         CALL  "FC071_CleaningPiston"
         ( IN_WithCP                := "DB704_MH_Value".Mixinghead[5].WithCleaningPiston,
           IN_Ana_CP_State          := #AnaCp_StatB,
           IN_SWUEnabled            := "DB619_State_MPart".SWU[1].SWU_released."05",
           IN_ButtonCPForward       := "DB123_MH_IO_Signals".MH[5].IN.MH_CP_forward,
           IN_ButtonCPback          := "DB123_MH_IO_Signals".MH[5].IN.MH_CP_backward,
           IN_CPForwardFromExternal := #Temp_CP_forward_external,
           IN_CPAfterShot           := "DB619_State_MPart".ShotMa[1].ShotData.CP_AfterShot,
           IN_PartshotDisabled      := "DB619_State_MPart".ShotMa[1].ShotData.ShotDisabled,
           IN_Blowing_OUT           := "DB614_MH_State".InertingMH[5].Start_Prepare_Purge_after_Shot,
           IN_CPProxSwitch          := "DB123_MH_IO_Signals".MH[5].IN.MH_APS_CleaningPiston,
           IN_SWUActive             := "DB619_State_MPart".SWU[1].Open_SWU_allone."05",
           IN_HydraulicOk           := "DB619_State_MPart".Machine[1].HydStartUp_finished,
           IN_ResetFaults           := "DB009_Faults".Faults_Reset_FKT_M1,
           IN_ControlVoltage        := "DB619_State_MPart".Operationmode[1].Controllvoltage,
           IN_OperatingModeValid    := "DB619_State_MPart".Operationmode[1].valid,
           IN_OperatingModeWithFoam := "DB619_State_MPart".Operationmode[1].Operation,
           IN_OperatingModeTestValv := "DB619_State_MPart".Operationmode[1].Test,
           IN_Lamptest              := "DB619_State_MPart".Operationmode[1].Lamptest,
           IN_ShotEnd               := "DB619_State_MPart".Cycle[1].PulsShotend,
           IN_FaultLevel_1          := "DB009_Faults".Fault_State_Grp_1_M1,
           IN_PressurizeTimeRunning := "DB619_State_MPart".Cycle[1].PressurizeTimeRuns,
           IN_ShotActive            := "DB619_State_MPart".Cycle[1].ShotRuns,
           IN_CycleRunning          := "DB619_State_MPart".Cycle[1].running,
           IN_RmpCtrlChangeTimeEnd  := "DB619_State_MPart".Cycle[1].RmpCtrlChangeTimeEnd,
           IN_StandbyTimeRunning    := "DB619_State_MPart".Cycle[1].StandByTimeRuns,
           IN_RmpCycleEnd           := "DB619_State_MPart".Cycle[1].PulseCycleEnd,
           IN_CPTimer               := "TM_RunTime_CP05",
           IN_TMCheckHomePos        := "TM_FltCPHomePos_CP05",
           Values                   := "DB704_MH_Value".Mixinghead[5].Cleaning_Piston,
           OUT_ValveCPForward       := "DB123_MH_IO_Signals".MH[5].OUT.MH.V_CP_Forward_MH,
           OUT_LampCPBack           := "DB123_MH_IO_Signals".MH[5].OUT.MH.H_CP_Back_MH,
           IO_CPIsOk                := "DB619_State_MPart".Mixinghead[1].Cleaningpiston_OK,
           IO_ReqHydrForCleaning    := "DB611_Hydraulic_State".MH_Hydraulic[1].Request_from_CP,
           IO_Status                := "DB614_MH_State".MH_CleaningPiston[5],
           IO_Fault                 := "DB824_Error_MH_CP".CPiston[5],
           IO_NewFault              := "DB009_Faults".Faultschanging_M1,
           IO_FaultLevel_1          := "DB009_Faults".Faults_FKT_Grp_1_M1,
           IO_FaultLevel_2          := "DB009_Faults".Faults_FKT_Grp_2_M1,
           IO_FaultLevel_3          := "DB009_Faults".Faults_FKT_Grp_3_M1
         );
END_REGION

REGION Network 11: Activate cleaning piston mixinghead by external signal
         A     "DB005_RS<->Extern".MC_Interface[6].Data_from_MC.CP_forward;
         =     #Temp_CP_forward_external;
END_REGION

REGION Network 12: Cleaning piston mixinghead 06
         CALL  BLKMOV
         ( SRCBLK  := "DB123_MH_IO_Signals".MH[6].IN.CleaningPistonState,
           RET_VAL := #RetValSFC,
           DSTBLK  := #AnaCp_Stat
         );

         L     #AnaCp_Stat;
         SRW   8;
         T     #AnaCp_StatB;

         CALL  "FC071_CleaningPiston"
         ( IN_WithCP                := "DB704_MH_Value".Mixinghead[6].WithCleaningPiston,
           IN_Ana_CP_State          := #AnaCp_StatB,
           IN_SWUEnabled            := "DB619_State_MPart".SWU[1].SWU_released."06",
           IN_ButtonCPForward       := "DB123_MH_IO_Signals".MH[6].IN.MH_CP_forward,
           IN_ButtonCPback          := "DB123_MH_IO_Signals".MH[6].IN.MH_CP_backward,
           IN_CPForwardFromExternal := #Temp_CP_forward_external,
           IN_CPAfterShot           := "DB619_State_MPart".ShotMa[1].ShotData.CP_AfterShot,
           IN_PartshotDisabled      := "DB619_State_MPart".ShotMa[1].ShotData.ShotDisabled,
           IN_Blowing_OUT           := "DB614_MH_State".InertingMH[6].Start_Prepare_Purge_after_Shot,
           IN_CPProxSwitch          := "DB123_MH_IO_Signals".MH[6].IN.MH_APS_CleaningPiston,
           IN_SWUActive             := "DB619_State_MPart".SWU[1].Open_SWU_allone."06",
           IN_HydraulicOk           := "DB619_State_MPart".Machine[1].HydStartUp_finished,
           IN_ResetFaults           := "DB009_Faults".Faults_Reset_FKT_M1,
           IN_ControlVoltage        := "DB619_State_MPart".Operationmode[1].Controllvoltage,
           IN_OperatingModeValid    := "DB619_State_MPart".Operationmode[1].valid,
           IN_OperatingModeWithFoam := "DB619_State_MPart".Operationmode[1].Operation,
           IN_OperatingModeTestValv := "DB619_State_MPart".Operationmode[1].Test,
           IN_Lamptest              := "DB619_State_MPart".Operationmode[1].Lamptest,
           IN_ShotEnd               := "DB619_State_MPart".Cycle[1].PulsShotend,
           IN_FaultLevel_1          := "DB009_Faults".Fault_State_Grp_1_M1,
           IN_PressurizeTimeRunning := "DB619_State_MPart".Cycle[1].PressurizeTimeRuns,
           IN_ShotActive            := "DB619_State_MPart".Cycle[1].ShotRuns,
           IN_CycleRunning          := "DB619_State_MPart".Cycle[1].running,
           IN_RmpCtrlChangeTimeEnd  := "DB619_State_MPart".Cycle[1].RmpCtrlChangeTimeEnd,
           IN_StandbyTimeRunning    := "DB619_State_MPart".Cycle[1].StandByTimeRuns,
           IN_RmpCycleEnd           := "DB619_State_MPart".Cycle[1].PulseCycleEnd,
           IN_CPTimer               := "TM_RunTime_CP06",
           IN_TMCheckHomePos        := "TM_FltCPHomePos_CP06",
           Values                   := "DB704_MH_Value".Mixinghead[6].Cleaning_Piston,
           OUT_ValveCPForward       := "DB123_MH_IO_Signals".MH[6].OUT.MH.V_CP_Forward_MH,
           OUT_LampCPBack           := "DB123_MH_IO_Signals".MH[6].OUT.MH.H_CP_Back_MH,
           IO_CPIsOk                := "DB619_State_MPart".Mixinghead[1].Cleaningpiston_OK,
           IO_ReqHydrForCleaning    := "DB611_Hydraulic_State".MH_Hydraulic[1].Request_from_CP,
           IO_Status                := "DB614_MH_State".MH_CleaningPiston[6],
           IO_Fault                 := "DB824_Error_MH_CP".CPiston[6],
           IO_NewFault              := "DB009_Faults".Faultschanging_M1,
           IO_FaultLevel_1          := "DB009_Faults".Faults_FKT_Grp_1_M1,
           IO_FaultLevel_2          := "DB009_Faults".Faults_FKT_Grp_2_M1,
           IO_FaultLevel_3          := "DB009_Faults".Faults_FKT_Grp_3_M1
         );
END_REGION

REGION Network 13: Activate cleaning piston mixinghead by external signal
         A     "DB005_RS<->Extern".MC_Interface[7].Data_from_MC.CP_forward;
         =     #Temp_CP_forward_external;
END_REGION

REGION Network 14: Cleaning piston mixinghead 07
         CALL  BLKMOV
         ( SRCBLK  := "DB123_MH_IO_Signals".MH[7].IN.CleaningPistonState,
           RET_VAL := #RetValSFC,
           DSTBLK  := #AnaCp_Stat
         );

         L     #AnaCp_Stat;
         SRW   8;
         T     #AnaCp_StatB;

         CALL  "FC071_CleaningPiston"
         ( IN_WithCP                := "DB704_MH_Value".Mixinghead[7].WithCleaningPiston,
           IN_Ana_CP_State          := #AnaCp_StatB,
           IN_SWUEnabled            := "DB619_State_MPart".SWU[1].SWU_released."07",
           IN_ButtonCPForward       := "DB123_MH_IO_Signals".MH[7].IN.MH_CP_forward,
           IN_ButtonCPback          := "DB123_MH_IO_Signals".MH[7].IN.MH_CP_backward,
           IN_CPForwardFromExternal := #Temp_CP_forward_external,
           IN_CPAfterShot           := "DB619_State_MPart".ShotMa[1].ShotData.CP_AfterShot,
           IN_PartshotDisabled      := "DB619_State_MPart".ShotMa[1].ShotData.ShotDisabled,
           IN_Blowing_OUT           := "DB614_MH_State".InertingMH[7].Start_Prepare_Purge_after_Shot,
           IN_CPProxSwitch          := "DB123_MH_IO_Signals".MH[7].IN.MH_APS_CleaningPiston,
           IN_SWUActive             := "DB619_State_MPart".SWU[1].Open_SWU_allone."07",
           IN_HydraulicOk           := "DB619_State_MPart".Machine[1].HydStartUp_finished,
           IN_ResetFaults           := "DB009_Faults".Faults_Reset_FKT_M1,
           IN_ControlVoltage        := "DB619_State_MPart".Operationmode[1].Controllvoltage,
           IN_OperatingModeValid    := "DB619_State_MPart".Operationmode[1].valid,
           IN_OperatingModeWithFoam := "DB619_State_MPart".Operationmode[1].Operation,
           IN_OperatingModeTestValv := "DB619_State_MPart".Operationmode[1].Test,
           IN_Lamptest              := "DB619_State_MPart".Operationmode[1].Lamptest,
           IN_ShotEnd               := "DB619_State_MPart".Cycle[1].PulsShotend,
           IN_FaultLevel_1          := "DB009_Faults".Fault_State_Grp_1_M1,
           IN_PressurizeTimeRunning := "DB619_State_MPart".Cycle[1].PressurizeTimeRuns,
           IN_ShotActive            := "DB619_State_MPart".Cycle[1].ShotRuns,
           IN_CycleRunning          := "DB619_State_MPart".Cycle[1].running,
           IN_RmpCtrlChangeTimeEnd  := "DB619_State_MPart".Cycle[1].RmpCtrlChangeTimeEnd,
           IN_StandbyTimeRunning    := "DB619_State_MPart".Cycle[1].StandByTimeRuns,
           IN_RmpCycleEnd           := "DB619_State_MPart".Cycle[1].PulseCycleEnd,
           IN_CPTimer               := "TM_RunTime_CP07",
           IN_TMCheckHomePos        := "TM_FltCPHomePos_CP07",
           Values                   := "DB704_MH_Value".Mixinghead[7].Cleaning_Piston,
           OUT_ValveCPForward       := "DB123_MH_IO_Signals".MH[7].OUT.MH.V_CP_Forward_MH,
           OUT_LampCPBack           := "DB123_MH_IO_Signals".MH[7].OUT.MH.H_CP_Back_MH,
           IO_CPIsOk                := "DB619_State_MPart".Mixinghead[1].Cleaningpiston_OK,
           IO_ReqHydrForCleaning    := "DB611_Hydraulic_State".MH_Hydraulic[1].Request_from_CP,
           IO_Status                := "DB614_MH_State".MH_CleaningPiston[7],
           IO_Fault                 := "DB824_Error_MH_CP".CPiston[7],
           IO_NewFault              := "DB009_Faults".Faultschanging_M1,
           IO_FaultLevel_1          := "DB009_Faults".Faults_FKT_Grp_1_M1,
           IO_FaultLevel_2          := "DB009_Faults".Faults_FKT_Grp_2_M1,
           IO_FaultLevel_3          := "DB009_Faults".Faults_FKT_Grp_3_M1
         );
END_REGION

REGION Network 15: Activate cleaning piston mixinghead by external signal
         A     "DB005_RS<->Extern".MC_Interface[8].Data_from_MC.CP_forward;
         =     #Temp_CP_forward_external;
END_REGION

REGION Network 16: Cleaning piston mixinghead 08
         CALL  BLKMOV
         ( SRCBLK  := "DB123_MH_IO_Signals".MH[8].IN.CleaningPistonState,
           RET_VAL := #RetValSFC,
           DSTBLK  := #AnaCp_Stat
         );

         L     #AnaCp_Stat;
         SRW   8;
         T     #AnaCp_StatB;

         CALL  "FC071_CleaningPiston"
         ( IN_WithCP                := "DB704_MH_Value".Mixinghead[8].WithCleaningPiston,
           IN_Ana_CP_State          := #AnaCp_StatB,
           IN_SWUEnabled            := "DB619_State_MPart".SWU[1].SWU_released."08",
           IN_ButtonCPForward       := "DB123_MH_IO_Signals".MH[8].IN.MH_CP_forward,
           IN_ButtonCPback          := "DB123_MH_IO_Signals".MH[8].IN.MH_CP_backward,
           IN_CPForwardFromExternal := #Temp_CP_forward_external,
           IN_CPAfterShot           := "DB619_State_MPart".ShotMa[1].ShotData.CP_AfterShot,
           IN_PartshotDisabled      := "DB619_State_MPart".ShotMa[1].ShotData.ShotDisabled,
           IN_Blowing_OUT           := "DB614_MH_State".InertingMH[8].Start_Prepare_Purge_after_Shot,
           IN_CPProxSwitch          := "DB123_MH_IO_Signals".MH[8].IN.MH_APS_CleaningPiston,
           IN_SWUActive             := "DB619_State_MPart".SWU[1].Open_SWU_allone."08",
           IN_HydraulicOk           := "DB619_State_MPart".Machine[1].HydStartUp_finished,
           IN_ResetFaults           := "DB009_Faults".Faults_Reset_FKT_M1,
           IN_ControlVoltage        := "DB619_State_MPart".Operationmode[1].Controllvoltage,
           IN_OperatingModeValid    := "DB619_State_MPart".Operationmode[1].valid,
           IN_OperatingModeWithFoam := "DB619_State_MPart".Operationmode[1].Operation,
           IN_OperatingModeTestValv := "DB619_State_MPart".Operationmode[1].Test,
           IN_Lamptest              := "DB619_State_MPart".Operationmode[1].Lamptest,
           IN_ShotEnd               := "DB619_State_MPart".Cycle[1].PulsShotend,
           IN_FaultLevel_1          := "DB009_Faults".Fault_State_Grp_1_M1,
           IN_PressurizeTimeRunning := "DB619_State_MPart".Cycle[1].PressurizeTimeRuns,
           IN_ShotActive            := "DB619_State_MPart".Cycle[1].ShotRuns,
           IN_CycleRunning          := "DB619_State_MPart".Cycle[1].running,
           IN_RmpCtrlChangeTimeEnd  := "DB619_State_MPart".Cycle[1].RmpCtrlChangeTimeEnd,
           IN_StandbyTimeRunning    := "DB619_State_MPart".Cycle[1].StandByTimeRuns,
           IN_RmpCycleEnd           := "DB619_State_MPart".Cycle[1].PulseCycleEnd,
           IN_CPTimer               := "TM_RunTime_CP08",
           IN_TMCheckHomePos        := "TM_FltCPHomePos_CP08",
           Values                   := "DB704_MH_Value".Mixinghead[8].Cleaning_Piston,
           OUT_ValveCPForward       := "DB123_MH_IO_Signals".MH[8].OUT.MH.V_CP_Forward_MH,
           OUT_LampCPBack           := "DB123_MH_IO_Signals".MH[8].OUT.MH.H_CP_Back_MH,
           IO_CPIsOk                := "DB619_State_MPart".Mixinghead[1].Cleaningpiston_OK,
           IO_ReqHydrForCleaning    := "DB611_Hydraulic_State".MH_Hydraulic[1].Request_from_CP,
           IO_Status                := "DB614_MH_State".MH_CleaningPiston[8],
           IO_Fault                 := "DB824_Error_MH_CP".CPiston[8],
           IO_NewFault              := "DB009_Faults".Faultschanging_M1,
           IO_FaultLevel_1          := "DB009_Faults".Faults_FKT_Grp_1_M1,
           IO_FaultLevel_2          := "DB009_Faults".Faults_FKT_Grp_2_M1,
           IO_FaultLevel_3          := "DB009_Faults".Faults_FKT_Grp_3_M1
         );
END_REGION

REGION Network 17: Activate cleaning piston mixinghead by external signal
         A     "DB005_RS<->Extern".MC_Interface[9].Data_from_MC.CP_forward;
         =     #Temp_CP_forward_external;
END_REGION

REGION Network 18: Cleaning piston mixinghead 09
         CALL  BLKMOV
         ( SRCBLK  := "DB123_MH_IO_Signals".MH[9].IN.CleaningPistonState,
           RET_VAL := #RetValSFC,
           DSTBLK  := #AnaCp_Stat
         );

         L     #AnaCp_Stat;
         SRW   8;
         T     #AnaCp_StatB;

         CALL  "FC071_CleaningPiston"
         ( IN_WithCP                := "DB704_MH_Value".Mixinghead[9].WithCleaningPiston,
           IN_Ana_CP_State          := #AnaCp_StatB,
           IN_SWUEnabled            := "DB619_State_MPart".SWU[1].SWU_released."09",
           IN_ButtonCPForward       := "DB123_MH_IO_Signals".MH[9].IN.MH_CP_forward,
           IN_ButtonCPback          := "DB123_MH_IO_Signals".MH[9].IN.MH_CP_backward,
           IN_CPForwardFromExternal := #Temp_CP_forward_external,
           IN_CPAfterShot           := "DB619_State_MPart".ShotMa[1].ShotData.CP_AfterShot,
           IN_PartshotDisabled      := "DB619_State_MPart".ShotMa[1].ShotData.ShotDisabled,
           IN_Blowing_OUT           := "DB614_MH_State".InertingMH[9].Start_Prepare_Purge_after_Shot,
           IN_CPProxSwitch          := "DB123_MH_IO_Signals".MH[9].IN.MH_APS_CleaningPiston,
           IN_SWUActive             := "DB619_State_MPart".SWU[1].Open_SWU_allone."09",
           IN_HydraulicOk           := "DB619_State_MPart".Machine[1].HydStartUp_finished,
           IN_ResetFaults           := "DB009_Faults".Faults_Reset_FKT_M1,
           IN_ControlVoltage        := "DB619_State_MPart".Operationmode[1].Controllvoltage,
           IN_OperatingModeValid    := "DB619_State_MPart".Operationmode[1].valid,
           IN_OperatingModeWithFoam := "DB619_State_MPart".Operationmode[1].Operation,
           IN_OperatingModeTestValv := "DB619_State_MPart".Operationmode[1].Test,
           IN_Lamptest              := "DB619_State_MPart".Operationmode[1].Lamptest,
           IN_ShotEnd               := "DB619_State_MPart".Cycle[1].PulsShotend,
           IN_FaultLevel_1          := "DB009_Faults".Fault_State_Grp_1_M1,
           IN_PressurizeTimeRunning := "DB619_State_MPart".Cycle[1].PressurizeTimeRuns,
           IN_ShotActive            := "DB619_State_MPart".Cycle[1].ShotRuns,
           IN_CycleRunning          := "DB619_State_MPart".Cycle[1].running,
           IN_RmpCtrlChangeTimeEnd  := "DB619_State_MPart".Cycle[1].RmpCtrlChangeTimeEnd,
           IN_StandbyTimeRunning    := "DB619_State_MPart".Cycle[1].StandByTimeRuns,
           IN_RmpCycleEnd           := "DB619_State_MPart".Cycle[1].PulseCycleEnd,
           IN_CPTimer               := "TM_RunTime_CP09",
           IN_TMCheckHomePos        := "TM_FltCPHomePos_CP09",
           Values                   := "DB704_MH_Value".Mixinghead[9].Cleaning_Piston,
           OUT_ValveCPForward       := "DB123_MH_IO_Signals".MH[9].OUT.MH.V_CP_Forward_MH,
           OUT_LampCPBack           := "DB123_MH_IO_Signals".MH[9].OUT.MH.H_CP_Back_MH,
           IO_CPIsOk                := "DB619_State_MPart".Mixinghead[1].Cleaningpiston_OK,
           IO_ReqHydrForCleaning    := "DB611_Hydraulic_State".MH_Hydraulic[1].Request_from_CP,
           IO_Status                := "DB614_MH_State".MH_CleaningPiston[9],
           IO_Fault                 := "DB824_Error_MH_CP".CPiston[9],
           IO_NewFault              := "DB009_Faults".Faultschanging_M1,
           IO_FaultLevel_1          := "DB009_Faults".Faults_FKT_Grp_1_M1,
           IO_FaultLevel_2          := "DB009_Faults".Faults_FKT_Grp_2_M1,
           IO_FaultLevel_3          := "DB009_Faults".Faults_FKT_Grp_3_M1
         );
END_REGION

REGION Network 19: Activate cleaning piston mixinghead by external signal
         A     "DB005_RS<->Extern".MC_Interface[10].Data_from_MC.CP_forward;
         =     #Temp_CP_forward_external;
END_REGION

REGION Network 20: Cleaning piston mixinghead 10
         CALL  BLKMOV
         ( SRCBLK  := "DB123_MH_IO_Signals".MH[10].IN.CleaningPistonState,
           RET_VAL := #RetValSFC,
           DSTBLK  := #AnaCp_Stat
         );

         L     #AnaCp_Stat;
         SRW   8;
         T     #AnaCp_StatB;

         CALL  "FC071_CleaningPiston"
         ( IN_WithCP                := "DB704_MH_Value".Mixinghead[10].WithCleaningPiston,
           IN_Ana_CP_State          := #AnaCp_StatB,
           IN_SWUEnabled            := "DB619_State_MPart".SWU[1].SWU_released."10",
           IN_ButtonCPForward       := "DB123_MH_IO_Signals".MH[10].IN.MH_CP_forward,
           IN_ButtonCPback          := "DB123_MH_IO_Signals".MH[10].IN.MH_CP_backward,
           IN_CPForwardFromExternal := #Temp_CP_forward_external,
           IN_CPAfterShot           := "DB619_State_MPart".ShotMa[1].ShotData.CP_AfterShot,
           IN_PartshotDisabled      := "DB619_State_MPart".ShotMa[1].ShotData.ShotDisabled,
           IN_Blowing_OUT           := "DB614_MH_State".InertingMH[10].Start_Prepare_Purge_after_Shot,
           IN_CPProxSwitch          := "DB123_MH_IO_Signals".MH[10].IN.MH_APS_CleaningPiston,
           IN_SWUActive             := "DB619_State_MPart".SWU[1].Open_SWU_allone."10",
           IN_HydraulicOk           := "DB619_State_MPart".Machine[1].HydStartUp_finished,
           IN_ResetFaults           := "DB009_Faults".Faults_Reset_FKT_M1,
           IN_ControlVoltage        := "DB619_State_MPart".Operationmode[1].Controllvoltage,
           IN_OperatingModeValid    := "DB619_State_MPart".Operationmode[1].valid,
           IN_OperatingModeWithFoam := "DB619_State_MPart".Operationmode[1].Operation,
           IN_OperatingModeTestValv := "DB619_State_MPart".Operationmode[1].Test,
           IN_Lamptest              := "DB619_State_MPart".Operationmode[1].Lamptest,
           IN_ShotEnd               := "DB619_State_MPart".Cycle[1].PulsShotend,
           IN_FaultLevel_1          := "DB009_Faults".Fault_State_Grp_1_M1,
           IN_PressurizeTimeRunning := "DB619_State_MPart".Cycle[1].PressurizeTimeRuns,
           IN_ShotActive            := "DB619_State_MPart".Cycle[1].ShotRuns,
           IN_CycleRunning          := "DB619_State_MPart".Cycle[1].running,
           IN_RmpCtrlChangeTimeEnd  := "DB619_State_MPart".Cycle[1].RmpCtrlChangeTimeEnd,
           IN_StandbyTimeRunning    := "DB619_State_MPart".Cycle[1].StandByTimeRuns,
           IN_RmpCycleEnd           := "DB619_State_MPart".Cycle[1].PulseCycleEnd,
           IN_CPTimer               := "TM_RunTime_CP10",
           IN_TMCheckHomePos        := "TM_FltCPHomePos_CP10",
           Values                   := "DB704_MH_Value".Mixinghead[10].Cleaning_Piston,
           OUT_ValveCPForward       := "DB123_MH_IO_Signals".MH[10].OUT.MH.V_CP_Forward_MH,
           OUT_LampCPBack           := "DB123_MH_IO_Signals".MH[10].OUT.MH.H_CP_Back_MH,
           IO_CPIsOk                := "DB619_State_MPart".Mixinghead[1].Cleaningpiston_OK,
           IO_ReqHydrForCleaning    := "DB611_Hydraulic_State".MH_Hydraulic[1].Request_from_CP,
           IO_Status                := "DB614_MH_State".MH_CleaningPiston[10],
           IO_Fault                 := "DB824_Error_MH_CP".CPiston[10],
           IO_NewFault              := "DB009_Faults".Faultschanging_M1,
           IO_FaultLevel_1          := "DB009_Faults".Faults_FKT_Grp_1_M1,
           IO_FaultLevel_2          := "DB009_Faults".Faults_FKT_Grp_2_M1,
           IO_FaultLevel_3          := "DB009_Faults".Faults_FKT_Grp_3_M1
         );
END_REGION

REGION Network 21: Reset request hydraulic from cleaning piston
         A     "DB611_Hydraulic_State".MH_Hydraulic[1].Request_from_CP;
         L     S5T#10S;
         SD    "TM_HydrForCPoffM1";

         A     "TM_HydrForCPoffM1";
         R     "DB611_Hydraulic_State".MH_Hydraulic[1].Request_from_CP;
END_REGION
END_FUNCTION_BLOCK

FUNCTION_BLOCK "FB019_FoamingCycle_M1"   // FB19, STL
TITLE = Foaming Cycle Control
{ S7_Optimized_Access := 'FALSE' }
AUTHOR : KT242
VERSION : 0.1
// Foaming Cycle Control
   VAR_TEMP
      Temp_MH_No : "UDT001_DWord_1_32";
      RetValSFC : Int;
      ProCanMH_State : Struct
         NoShotReleaseFromCP : Bool;   // No Shot Release from Cleaning Piston
         NoShotReleaseFromExtern : Bool;   // No Shot Release from Extern
         Ready4Shot : Bool;   // Ready for Shot
         shotactive_MH : Bool;   // Shot is active
         shotdone_MH : Bool;   // Shot finished
         Spare5 : Bool;
         Spare6 : Bool;
         Spare7 : Bool;
         SPFopening_MH : Bool;   // Steering piston fault opening time exceeded
         SPFclosing_MH : Bool;   // Steering piston fault closing time exceeded
         SPFopen_MH : Bool;   // Steering piston fault MH is open before shot
         SPFclosed_MH : Bool;   // Steering piston MH closed before end of shot
         MHBouncing : Bool;   // Partner has shot enabled
         SPFaborted_SoftwareRelease : Bool;
         SPFaborted_CP : Bool;
         SPFabortet_HardwareRelease : Bool;
      END_STRUCT;
      CycleRelease : Bool;
      Release_PBT1 : Bool;   // Release of pressure build up time
      ShotRunning : Bool;
      StartCycle : Bool;
      CtrlChangeTime : S5Time;
   END_VAR
BEGIN

REGION Network 1: Release foaming cycle
         A     "DB619_State_MPart".Operationmode[1].Auto;
         A     "DB619_State_MPart".Operationmode[1].Active;
         =     #CycleRelease;
END_REGION

REGION Network 2: Realease pressure build up (KLZ 1)
         A(;
         O     "DB110_Interf_Program_M1".Status_IF[1].IF_is_on_1_Position;
         O     "DB110_Interf_Program_M1".Status_IF[2].IF_is_on_1_Position;
         O     "DB110_Interf_Program_M1".Status_IF[3].IF_is_on_1_Position;
         O     "DB110_Interf_Program_M1".Status_IF[4].IF_is_on_1_Position;
         O     "DB110_Interf_Program_M1".Status_IF[5].IF_is_on_1_Position;
         O     "DB110_Interf_Program_M1".Status_IF[6].IF_is_on_1_Position;
         O     "DB110_Interf_Program_M1".Status_IF[7].IF_is_on_1_Position;
         O     "DB110_Interf_Program_M1".Status_IF[8].IF_is_on_1_Position;
         O     "DB110_Interf_Program_M1".Status_IF[9].IF_is_on_1_Position;
         O     "DB110_Interf_Program_M1".Status_IF[10].IF_is_on_1_Position;
         O     "DB110_Interf_Program_M1".Status_IF[11].IF_is_on_1_Position;
         O     "DB110_Interf_Program_M1".Status_IF[12].IF_is_on_1_Position;
         O     "DB619_State_MPart".Operationmode[1].Test;
         );
         AN    "DB619_State_MPart".SWU[1].Switchingtime_runs;
         A     "DB619_State_MPart".Cycle[1].running;
         AN    "TM_SwitchOnDelayFCPump";
         =     #Release_PBT1;
END_REGION

REGION Network 3: Modul indicates shot during production and service mode
         O     "DB123_MH_IO_Signals".MH[1].IN.MH_Status.shotactive_MH;
         O     "DB123_MH_IO_Signals".MH[2].IN.MH_Status.shotactive_MH;
         O     "DB123_MH_IO_Signals".MH[3].IN.MH_Status.shotactive_MH;
         O     "DB123_MH_IO_Signals".MH[4].IN.MH_Status.shotactive_MH;
         O     "DB123_MH_IO_Signals".MH[5].IN.MH_Status.shotactive_MH;
         O     "DB123_MH_IO_Signals".MH[6].IN.MH_Status.shotactive_MH;
         O     "DB123_MH_IO_Signals".MH[7].IN.MH_Status.shotactive_MH;
         O     "DB123_MH_IO_Signals".MH[8].IN.MH_Status.shotactive_MH;
         O     "DB123_MH_IO_Signals".MH[9].IN.MH_Status.shotactive_MH;
         O     "DB123_MH_IO_Signals".MH[10].IN.MH_Status.shotactive_MH;
         O     "DB123_MH_IO_Signals".MH[11].IN.MH_Status.shotactive_MH;
         O     "DB123_MH_IO_Signals".MH[12].IN.MH_Status.shotactive_MH;
         =     #ShotRunning;
         =     "M_ShotActive";
END_REGION

REGION Network 4
         A     "DB619_State_MPart".ToolMa[1].ShotFound;
         AN    "DB619_State_MPart".Cycle[1].PulsShotend;
         A     "DB619_State_MPart".ToolMa[1].Tool.EnableTool;
         =     #StartCycle;
END_REGION

REGION Network 5: Sequence of foamingcycle with all steps and timers
   // At the end of the shot, the actual MH number is stored in MW201
         A     "DB619_State_MPart".Cycle[1].PulsShotend;
         JCN   noShEnd;

         L     "DB619_State_MPart".ShotMa[1].ShotData.MH_No;
         T     "PulsShotend_M1_MH_No";

   noShEnd:NOP   0;

   // When the next shot is recognized, the actual MH number is stored in MW212
         A     "DB619_State_MPart".ToolMa[1].ShotFound;
         FP    "HM_FP_ShotFound_M1";
         JCN   noShFnd;

         L     "DB619_State_MPart".ShotMa[1].ShotData.MH_No;
         T     "NextShot_M1_MH_No";

   noShFnd:NOP   0;

   // If MW201 and MW212 are different, the control changing time is longer
         AN(;
         L     "PulsShotend_M1_MH_No";
         L     "NextShot_M1_MH_No";
         ==I;
         );
         JC    LongT;

   // If MW201 and MW212 are equal, the control changing time is shorter
         JU    ShortT;

   LongT:L     "DB700_Machine".Machine[1].CtrlChangeTime2;
         T     #CtrlChangeTime;
         JU    end1;

   ShortT:L     "DB700_Machine".Machine[1].CtrlChangeTime1;
         T     #CtrlChangeTime;

   end1: NOP   0;


         CALL  "FC091_PouringCycle"
         ( IN_OMAutomatic          := "DB619_State_MPart".Operationmode[1].Auto,
           IN_OMChange             := "DB619_State_MPart".Operationmode[1].Edge_OM_Change,
           IN_ResetFaults          := "DB009_Faults".Faults_Reset_FKT_M1,
           IN_LampTest             := "DB619_State_MPart".Operationmode[1].Lamptest,
           IN_EnableCycle          := #CycleRelease,
           IN_EnablePressurizeTime := #Release_PBT1,
           IN_ShotActive           := #ShotRunning,
           IN_Hydraulics_OK        := "DB619_State_MPart".Machine[1].HydStartUp_finished,
           IN_DW_PressurizeTime    := "DB700_Machine".Machine[1].PressureBuildUpTime,
           IN_DW_StandByTime       := "DB700_Machine".Machine[1].StandByTime,
           IN_DW_CntrlChangeTime   := #CtrlChangeTime,  //"DB700_Machine".Machine[1].CtrlChangeTime1
           IN_DW_MaxWaitTime       := "DB700_Machine".Machine[1].Max_WaitTime,
           IN_DW_MaxShotTime       := "DB700_Machine".Machine[1].Max_ShotTime,
           IN_Cycletimer           := "TM_CycleTimer_M1",
           IN_FaultLevel_1         := "DB009_Faults".Fault_State_Grp_1_M1,
           IN_FaultLevel_2         := "DB009_Faults".Fault_State_Grp_2_M1,
           OUT_LampMachineOK       := "H_Ready_for_Operation_M1",
           IO_Status               := "DB619_State_MPart".Cycle[1],
           IO_Fault                := "DB829_Error_Machine".PouringCycle[1],
           IO_FaultLevel_1         := "DB009_Faults".Faults_FKT_Grp_1_M1,
           IO_FaultLevel_2         := "DB009_Faults".Faults_FKT_Grp_2_M1,
           IO_FaultLevel_3         := "DB009_Faults".Faults_FKT_Grp_3_M1,
           IO_NewFault             := "DB009_Faults".Faultschanging_M1,
           IO_StartShotCycle       := #StartCycle,
           IO_StopShotCycle        := "DB110_Interf_Program_M1".Bits.Stop_Cycle  // "DB610_State_MPart".ShotSelMa[1].StopCycle
         );


   //--------------------------------------------------------------------------------
   //    State shot:
   //               ShotState: Value 0 -> Shot OK
   //                          Value  1  Array[0] ->  1 - Shot stopped by error
   //                          Value  2  Array[1] ->  1 - Shot stopped by break
   //                          Value  4  Array[2] ->  1 - Operation; 0 - Service Shot
   //                          Value  8  Array[3] ->  1 - Mixinghead at manual mode
   //--------------------------------------------------------------------------------
         A     #ShotRunning;
         FP    "HF_FP_ShotRunning";
         R     "DB919_ShotResultMach".ShotResult_Ma[1].General.ShotState[0];
         R     "DB919_ShotResultMach".ShotResult_Ma[1].General.ShotState[1];
         R     "DB919_ShotResultMach".ShotResult_Ma[1].General.ShotState[2];
         R     "DB919_ShotResultMach".ShotResult_Ma[1].General.ShotState[3];
         R     "DB919_ShotResultMach".ShotResult_Ma[1].General.ShotState[4];
         R     "ShotDisabledDuringShot";

         A     "DB619_State_MPart".ShotMa[1].ShotData.ShotDisabled;
         A     #ShotRunning;
         FP    "HF_ShotDisabledDuringShot";
         S     "ShotDisabledDuringShot";

         A     #ShotRunning;
         A     "DB009_Faults".Fault_State_Grp_1_M1;
         S     "DB919_ShotResultMach".ShotResult_Ma[1].General.ShotState[0];

         A     #ShotRunning;
         A     "DB110_Interf_Program_M1".Bits.Stop_Cycle;
         S     "DB919_ShotResultMach".ShotResult_Ma[1].General.ShotState[1];

         O     "ShotDisabledDuringShot";
         ON    "DB619_State_MPart".Operationmode[1].Operation;
         S     "DB919_ShotResultMach".ShotResult_Ma[1].General.ShotState[2];

   //-----------------------------------------------------------------------
   // MH at shot in manual mode at machine 1
   //-----------------------------------------------------------------------
         O(;
         A     "DB619_State_MPart".SWU[1].Open_SWU_allone."01";
         A     "DB123_MH_IO_Signals".MH[1].IN.MH_Manual_Mode;
         A     "DB619_State_MPart".MH_at_Machine[1]."01";
         );
         O(;
         A     "DB619_State_MPart".SWU[1].Open_SWU_allone."02";
         A     "DB123_MH_IO_Signals".MH[2].IN.MH_Manual_Mode;
         A     "DB619_State_MPart".MH_at_Machine[1]."02";
         );
         O(;
         A     "DB619_State_MPart".SWU[1].Open_SWU_allone."03";
         A     "DB123_MH_IO_Signals".MH[3].IN.MH_Manual_Mode;
         A     "DB619_State_MPart".MH_at_Machine[1]."03";
         );
         O(;
         A     "DB619_State_MPart".SWU[1].Open_SWU_allone."04";
         A     "DB123_MH_IO_Signals".MH[4].IN.MH_Manual_Mode;
         A     "DB619_State_MPart".MH_at_Machine[1]."04";
         );
         O(;
         A     "DB619_State_MPart".SWU[1].Open_SWU_allone."05";
         A     "DB123_MH_IO_Signals".MH[5].IN.MH_Manual_Mode;
         A     "DB619_State_MPart".MH_at_Machine[1]."05";
         );
         O(;
         A     "DB619_State_MPart".SWU[1].Open_SWU_allone."06";
         A     "DB123_MH_IO_Signals".MH[6].IN.MH_Manual_Mode;
         A     "DB619_State_MPart".MH_at_Machine[1]."06";
         );
         O(;
         A     "DB619_State_MPart".SWU[1].Open_SWU_allone."07";
         A     "DB123_MH_IO_Signals".MH[7].IN.MH_Manual_Mode;
         A     "DB619_State_MPart".MH_at_Machine[1]."07";
         );
         O(;
         A     "DB619_State_MPart".SWU[1].Open_SWU_allone."08";
         A     "DB123_MH_IO_Signals".MH[8].IN.MH_Manual_Mode;
         A     "DB619_State_MPart".MH_at_Machine[1]."08";
         );
         O(;
         A     "DB619_State_MPart".SWU[1].Open_SWU_allone."09";
         A     "DB123_MH_IO_Signals".MH[9].IN.MH_Manual_Mode;
         A     "DB619_State_MPart".MH_at_Machine[1]."09";
         );
         O(;
         A     "DB619_State_MPart".SWU[1].Open_SWU_allone."10";
         A     "DB123_MH_IO_Signals".MH[10].IN.MH_Manual_Mode;
         A     "DB619_State_MPart".MH_at_Machine[1]."10";
         );
         O(;
         A     "DB619_State_MPart".SWU[1].Open_SWU_allone."11";
         A     "DB123_MH_IO_Signals".MH[11].IN.MH_Manual_Mode;
         A     "DB619_State_MPart".MH_at_Machine[1]."11";
         );
         O(;
         A     "DB619_State_MPart".SWU[1].Open_SWU_allone."12";
         A     "DB123_MH_IO_Signals".MH[12].IN.MH_Manual_Mode;
         A     "DB619_State_MPart".MH_at_Machine[1]."12";
         );
         A     "DB619_State_MPart".Cycle[1].running;
         S     "DB919_ShotResultMach".ShotResult_Ma[1].General.ShotState[3];
END_REGION

REGION Network 6: Faults foaming cycle mixinghead 1 ... x
   // Mixinghead 1
         CALL  BLKMOV
         ( SRCBLK  := "DB123_MH_IO_Signals".MH[1].IN.MH_Status,
           RET_VAL := #RetValSFC,
           DSTBLK  := #ProCanMH_State
         );

         CALL  "FC096_Faults_MH"
         ( IN_ProCanMH_State     := #ProCanMH_State,  // ProCan-MH_Status MH01
           IN_Reset_Fault        := "DB009_Faults".Faults_Reset_FKT_M1,
           IN_CheckMH_Shot       := TRUE,
           IO_Any_ShotCycleState := "DB619_State_MPart".Cycle[1],
           IO_Any_MH_Fault       := "DB824_Error_MH_CP".MH_Control[1],
           IO_FaultLevel1        := "DB009_Faults".Faults_FKT_Grp_1_M1,
           IO_FaultLevel2        := "DB009_Faults".Faults_FKT_Grp_2_M1,
           IO_FaultLevel3        := "DB009_Faults".Faults_FKT_Grp_3_M1,
           IO_NewFault           := "DB009_Faults".Faultschanging_M1
         );

   // Mixinghead 2
         CALL  BLKMOV
         ( SRCBLK  := "DB123_MH_IO_Signals".MH[2].IN.MH_Status,
           RET_VAL := #RetValSFC,
           DSTBLK  := #ProCanMH_State
         );

         CALL  "FC096_Faults_MH"
         ( IN_ProCanMH_State     := #ProCanMH_State,  // ProCan-MH_Status MH02
           IN_Reset_Fault        := "DB009_Faults".Faults_Reset_FKT_M1,
           IN_CheckMH_Shot       := TRUE,
           IO_Any_ShotCycleState := "DB619_State_MPart".Cycle[1],
           IO_Any_MH_Fault       := "DB824_Error_MH_CP".MH_Control[2],
           IO_FaultLevel1        := "DB009_Faults".Faults_FKT_Grp_1_M1,
           IO_FaultLevel2        := "DB009_Faults".Faults_FKT_Grp_2_M1,
           IO_FaultLevel3        := "DB009_Faults".Faults_FKT_Grp_3_M1,
           IO_NewFault           := "DB009_Faults".Faultschanging_M1
         );

   // Mixinghead 3
         CALL  BLKMOV
         ( SRCBLK  := "DB123_MH_IO_Signals".MH[3].IN.MH_Status,
           RET_VAL := #RetValSFC,
           DSTBLK  := #ProCanMH_State
         );

         CALL  "FC096_Faults_MH"
         ( IN_ProCanMH_State     := #ProCanMH_State,  // ProCan-MH_Status MH03
           IN_Reset_Fault        := "DB009_Faults".Faults_Reset_FKT_M1,
           IN_CheckMH_Shot       := TRUE,
           IO_Any_ShotCycleState := "DB619_State_MPart".Cycle[1],
           IO_Any_MH_Fault       := "DB824_Error_MH_CP".MH_Control[3],
           IO_FaultLevel1        := "DB009_Faults".Faults_FKT_Grp_1_M1,
           IO_FaultLevel2        := "DB009_Faults".Faults_FKT_Grp_2_M1,
           IO_FaultLevel3        := "DB009_Faults".Faults_FKT_Grp_3_M1,
           IO_NewFault           := "DB009_Faults".Faultschanging_M1
         );

   // Mixinghead 4
         CALL  BLKMOV
         ( SRCBLK  := "DB123_MH_IO_Signals".MH[4].IN.MH_Status,
           RET_VAL := #RetValSFC,
           DSTBLK  := #ProCanMH_State
         );

         CALL  "FC096_Faults_MH"
         ( IN_ProCanMH_State     := #ProCanMH_State,  // ProCan-MH_Status MH04
           IN_Reset_Fault        := "DB009_Faults".Faults_Reset_FKT_M1,
           IN_CheckMH_Shot       := TRUE,
           IO_Any_ShotCycleState := "DB619_State_MPart".Cycle[1],
           IO_Any_MH_Fault       := "DB824_Error_MH_CP".MH_Control[4],
           IO_FaultLevel1        := "DB009_Faults".Faults_FKT_Grp_1_M1,
           IO_FaultLevel2        := "DB009_Faults".Faults_FKT_Grp_2_M1,
           IO_FaultLevel3        := "DB009_Faults".Faults_FKT_Grp_3_M1,
           IO_NewFault           := "DB009_Faults".Faultschanging_M1
         );

   // Mixinghead 5
         CALL  BLKMOV
         ( SRCBLK  := "DB123_MH_IO_Signals".MH[5].IN.MH_Status,
           RET_VAL := #RetValSFC,
           DSTBLK  := #ProCanMH_State
         );

         CALL  "FC096_Faults_MH"
         ( IN_ProCanMH_State     := #ProCanMH_State,  // ProCan-MH_Status MH05
           IN_Reset_Fault        := "DB009_Faults".Faults_Reset_FKT_M1,
           IN_CheckMH_Shot       := TRUE,
           IO_Any_ShotCycleState := "DB619_State_MPart".Cycle[1],
           IO_Any_MH_Fault       := "DB824_Error_MH_CP".MH_Control[5],
           IO_FaultLevel1        := "DB009_Faults".Faults_FKT_Grp_1_M1,
           IO_FaultLevel2        := "DB009_Faults".Faults_FKT_Grp_2_M1,
           IO_FaultLevel3        := "DB009_Faults".Faults_FKT_Grp_3_M1,
           IO_NewFault           := "DB009_Faults".Faultschanging_M1
         );

   // Mixinghead 6
         CALL  BLKMOV
         ( SRCBLK  := "DB123_MH_IO_Signals".MH[6].IN.MH_Status,
           RET_VAL := #RetValSFC,
           DSTBLK  := #ProCanMH_State
         );

         CALL  "FC096_Faults_MH"
         ( IN_ProCanMH_State     := #ProCanMH_State,  // ProCan-MH_Status MH06
           IN_Reset_Fault        := "DB009_Faults".Faults_Reset_FKT_M1,
           IN_CheckMH_Shot       := TRUE,
           IO_Any_ShotCycleState := "DB619_State_MPart".Cycle[1],
           IO_Any_MH_Fault       := "DB824_Error_MH_CP".MH_Control[6],
           IO_FaultLevel1        := "DB009_Faults".Faults_FKT_Grp_1_M1,
           IO_FaultLevel2        := "DB009_Faults".Faults_FKT_Grp_2_M1,
           IO_FaultLevel3        := "DB009_Faults".Faults_FKT_Grp_3_M1,
           IO_NewFault           := "DB009_Faults".Faultschanging_M1
         );

   // Mixinghead 7
         CALL  BLKMOV
         ( SRCBLK  := "DB123_MH_IO_Signals".MH[7].IN.MH_Status,
           RET_VAL := #RetValSFC,
           DSTBLK  := #ProCanMH_State
         );

         CALL  "FC096_Faults_MH"
         ( IN_ProCanMH_State     := #ProCanMH_State,  // ProCan-MH_Status MH07
           IN_Reset_Fault        := "DB009_Faults".Faults_Reset_FKT_M1,
           IN_CheckMH_Shot       := TRUE,
           IO_Any_ShotCycleState := "DB619_State_MPart".Cycle[1],
           IO_Any_MH_Fault       := "DB824_Error_MH_CP".MH_Control[7],
           IO_FaultLevel1        := "DB009_Faults".Faults_FKT_Grp_1_M1,
           IO_FaultLevel2        := "DB009_Faults".Faults_FKT_Grp_2_M1,
           IO_FaultLevel3        := "DB009_Faults".Faults_FKT_Grp_3_M1,
           IO_NewFault           := "DB009_Faults".Faultschanging_M1
         );

   // Mixinghead 8
         CALL  BLKMOV
         ( SRCBLK  := "DB123_MH_IO_Signals".MH[8].IN.MH_Status,
           RET_VAL := #RetValSFC,
           DSTBLK  := #ProCanMH_State
         );

         CALL  "FC096_Faults_MH"
         ( IN_ProCanMH_State     := #ProCanMH_State,  // ProCan-MH_Status MH08
           IN_Reset_Fault        := "DB009_Faults".Faults_Reset_FKT_M1,
           IN_CheckMH_Shot       := TRUE,
           IO_Any_ShotCycleState := "DB619_State_MPart".Cycle[1],
           IO_Any_MH_Fault       := "DB824_Error_MH_CP".MH_Control[8],
           IO_FaultLevel1        := "DB009_Faults".Faults_FKT_Grp_1_M1,
           IO_FaultLevel2        := "DB009_Faults".Faults_FKT_Grp_2_M1,
           IO_FaultLevel3        := "DB009_Faults".Faults_FKT_Grp_3_M1,
           IO_NewFault           := "DB009_Faults".Faultschanging_M1
         );

   // Mixinghead 9
         CALL  BLKMOV
         ( SRCBLK  := "DB123_MH_IO_Signals".MH[9].IN.MH_Status,
           RET_VAL := #RetValSFC,
           DSTBLK  := #ProCanMH_State
         );

         CALL  "FC096_Faults_MH"
         ( IN_ProCanMH_State     := #ProCanMH_State,  // ProCan-MH_Status MH09
           IN_Reset_Fault        := "DB009_Faults".Faults_Reset_FKT_M1,
           IN_CheckMH_Shot       := TRUE,
           IO_Any_ShotCycleState := "DB619_State_MPart".Cycle[1],
           IO_Any_MH_Fault       := "DB824_Error_MH_CP".MH_Control[9],
           IO_FaultLevel1        := "DB009_Faults".Faults_FKT_Grp_1_M1,
           IO_FaultLevel2        := "DB009_Faults".Faults_FKT_Grp_2_M1,
           IO_FaultLevel3        := "DB009_Faults".Faults_FKT_Grp_3_M1,
           IO_NewFault           := "DB009_Faults".Faultschanging_M1
         );

   // Mixinghead 10
         CALL  BLKMOV
         ( SRCBLK  := "DB123_MH_IO_Signals".MH[10].IN.MH_Status,
           RET_VAL := #RetValSFC,
           DSTBLK  := #ProCanMH_State
         );

         CALL  "FC096_Faults_MH"
         ( IN_ProCanMH_State     := #ProCanMH_State,  // ProCan-MH_Status MH10
           IN_Reset_Fault        := "DB009_Faults".Faults_Reset_FKT_M1,
           IN_CheckMH_Shot       := TRUE,
           IO_Any_ShotCycleState := "DB619_State_MPart".Cycle[1],
           IO_Any_MH_Fault       := "DB824_Error_MH_CP".MH_Control[10],
           IO_FaultLevel1        := "DB009_Faults".Faults_FKT_Grp_1_M1,
           IO_FaultLevel2        := "DB009_Faults".Faults_FKT_Grp_2_M1,
           IO_FaultLevel3        := "DB009_Faults".Faults_FKT_Grp_3_M1,
           IO_NewFault           := "DB009_Faults".Faultschanging_M1
         );

   // Mixinghead 11
         CALL  BLKMOV
         ( SRCBLK  := "DB123_MH_IO_Signals".MH[11].IN.MH_Status,
           RET_VAL := #RetValSFC,
           DSTBLK  := #ProCanMH_State
         );

         CALL  "FC096_Faults_MH"
         ( IN_ProCanMH_State     := #ProCanMH_State,  // ProCan-MH_Status MH11
           IN_Reset_Fault        := "DB009_Faults".Faults_Reset_FKT_M1,
           IN_CheckMH_Shot       := TRUE,
           IO_Any_ShotCycleState := "DB619_State_MPart".Cycle[1],
           IO_Any_MH_Fault       := "DB824_Error_MH_CP".MH_Control[11],
           IO_FaultLevel1        := "DB009_Faults".Faults_FKT_Grp_1_M1,
           IO_FaultLevel2        := "DB009_Faults".Faults_FKT_Grp_2_M1,
           IO_FaultLevel3        := "DB009_Faults".Faults_FKT_Grp_3_M1,
           IO_NewFault           := "DB009_Faults".Faultschanging_M1
         );

   // Mixinghead 12
         CALL  BLKMOV
         ( SRCBLK  := "DB123_MH_IO_Signals".MH[12].IN.MH_Status,
           RET_VAL := #RetValSFC,
           DSTBLK  := #ProCanMH_State
         );

         CALL  "FC096_Faults_MH"
         ( IN_ProCanMH_State     := #ProCanMH_State,  // ProCan-MH_Status MH12
           IN_Reset_Fault        := "DB009_Faults".Faults_Reset_FKT_M1,
           IN_CheckMH_Shot       := TRUE,
           IO_Any_ShotCycleState := "DB619_State_MPart".Cycle[1],
           IO_Any_MH_Fault       := "DB824_Error_MH_CP".MH_Control[12],
           IO_FaultLevel1        := "DB009_Faults".Faults_FKT_Grp_1_M1,
           IO_FaultLevel2        := "DB009_Faults".Faults_FKT_Grp_2_M1,
           IO_FaultLevel3        := "DB009_Faults".Faults_FKT_Grp_3_M1,
           IO_NewFault           := "DB009_Faults".Faultschanging_M1
         );
END_REGION

REGION Network 7
   //    CALL  "FC5029_InterfaceMouldProgram"
         CALL  "FC5030_InterfaceactualMHValue"
         ( IN_MachineNo := 1
         );
         CALL  "FC5031_InterfaceMachineGeneral";
         CALL  "FC5032_Last10Shot"
         ( IN_MachineNo := 1
         );
END_REGION
END_FUNCTION_BLOCK

FUNCTION_BLOCK "FB030_BallufReader"   // FB30, STL
TITLE = Schreib-/ Lesebaustein für Balluff Codeträgersystem (V1.8)
{ S7_Optimized_Access := 'FALSE' }
AUTHOR : Serrano
FAMILY : Ident
NAME : BIS60X2